(* Logix 5000 project; controller MV vendor 1 type 14 code 217 rev 31.11; software revision 31.00; part 23 of 53 *)
(* tags used below, declared in another part *)
   CheckTimeMask : INT;
   CWD : CHECKWORD_FLAGS;
   Delphi_Does_Eng_Func : BOOL;
   MC_CIP_AV01 : PlantItem;   // CIP_AV01
   MC_CIP_AV02 : PlantItem;   // CIP_AV02
   MC_CIP_AV05 : PlantItem;   // CIP_AV05
   MC_CIP_AV06 : PlantItem;   // CIP_AV06
   MC_CIP_AV07 : PlantItem;   // CIP_AV07
   MC_CIP_AV08 : PlantItem;   // CIP_AV08
   MC_CIP_AV09 : PlantItem;   // CIP_AV09
   MC_CIP_AV10 : PlantItem;   // CIP_AV10
   MC_N255 : INT[255];   // CHECKWORDS Plant item checkword s
   MC_R3R_DR : PlantItem;   // R3R_DR
   MC_R3S_DR : PlantItem;   // R3S_DR
   MC_R3V1 : PlantItem;   // R3V1
   MC_R3V2 : PlantItem;   // R3V2
   MC_SPV5 : PlantItem;   // SPV5
   TempChecktime : DINT;
(* MC_Common, continued *)

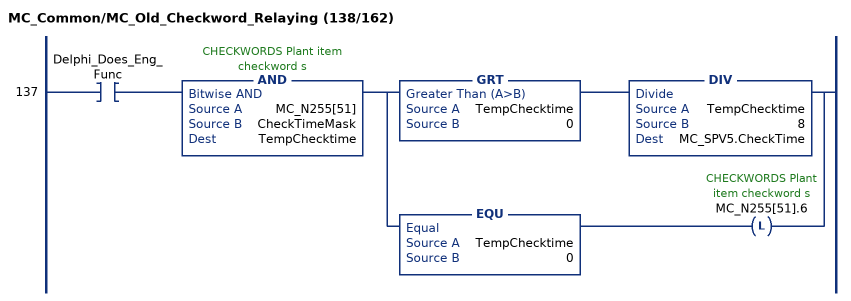
   [picture p410: MC_Common/MC_Old_Checkword_Relaying rungs 137-137]
   137: XIC(Delphi_Does_Eng_Func)AND(MC_N255[51],CheckTimeMask,TempChecktime)[GRT(TempChecktime,0) DIV(TempChecktime,8,MC_SPV5.CheckTime) ,EQU(TempChecktime,0) OTL(MC_N255[51].6) ];
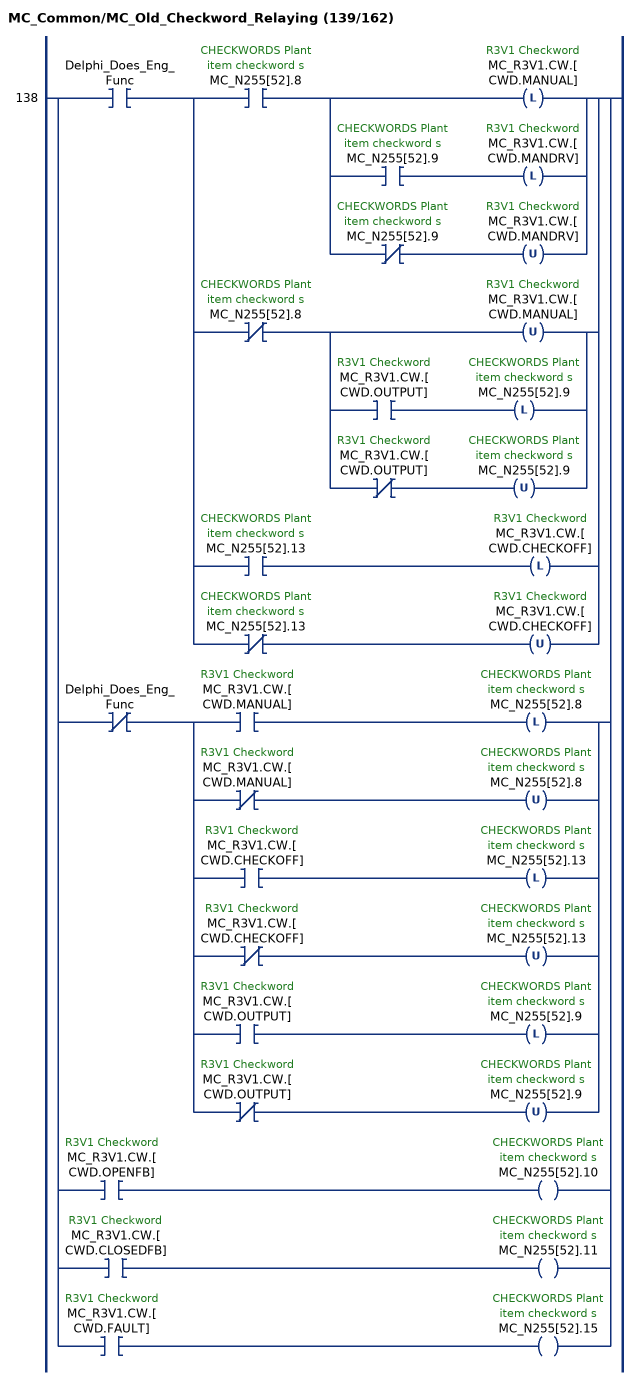
   138: [XIC(Delphi_Does_Eng_Func) [[XIC(MC_N255[52].8) [OTL(MC_R3V1.CW.[CWD.MANUAL]) ,XIC(MC_N255[52].9) OTL(MC_R3V1.CW.[CWD.MANDRV]) ,XIO(MC_N255[52].9) OTU(MC_R3V1.CW.[CWD.MANDRV]) ] ,XIO(MC_N255[52].8) [OTU(MC_R3V1.CW.[CWD.MANUAL]) ,[XIC(MC_R3V1.CW.[CWD.OUTPUT]) OTL(MC_N255[52].9) ,XIO(MC_R3V1.CW.[CWD.OUTPUT]) OTU(MC_N255[52].9) ] ] ] ,[XIC(MC_N255[52].13) OTL(MC_R3V1.CW.[CWD.CHECKOFF]) ,XIO(MC_N255[52].13) OTU(MC_R3V1.CW.[CWD.CHECKOFF]) ] ] ,XIO(Delphi_Does_Eng_Func) [[XIC(MC_R3V1.CW.[CWD.MANUAL]) OTL(MC_N255[52].8) ,XIO(MC_R3V1.CW.[CWD.MANUAL]) OTU(MC_N255[52].8) ] ,[XIC(MC_R3V1.CW.[CWD.CHECKOFF]) OTL(MC_N255[52].13) ,XIO(MC_R3V1.CW.[CWD.CHECKOFF]) OTU(MC_N255[52].13) ] ,[XIC(MC_R3V1.CW.[CWD.OUTPUT]) OTL(MC_N255[52].9) ,XIO(MC_R3V1.CW.[CWD.OUTPUT]) OTU(MC_N255[52].9) ] ] ,XIC(MC_R3V1.CW.[CWD.OPENFB]) OTE(MC_N255[52].10) ,XIC(MC_R3V1.CW.[CWD.CLOSEDFB]) OTE(MC_N255[52].11) ,XIC(MC_R3V1.CW.[CWD.FAULT]) OTE(MC_N255[52].15) ];
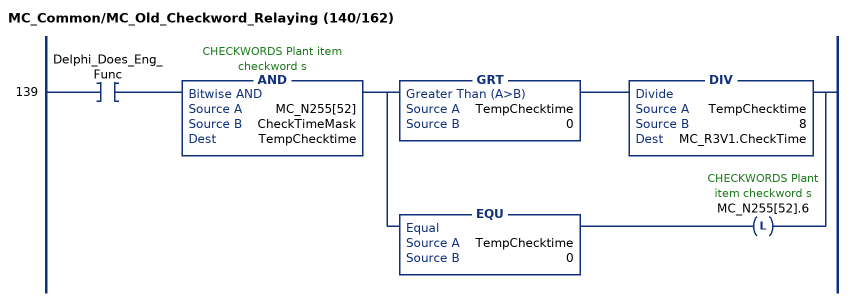
   139: XIC(Delphi_Does_Eng_Func)AND(MC_N255[52],CheckTimeMask,TempChecktime)[GRT(TempChecktime,0) DIV(TempChecktime,8,MC_R3V1.CheckTime) ,EQU(TempChecktime,0) OTL(MC_N255[52].6) ];
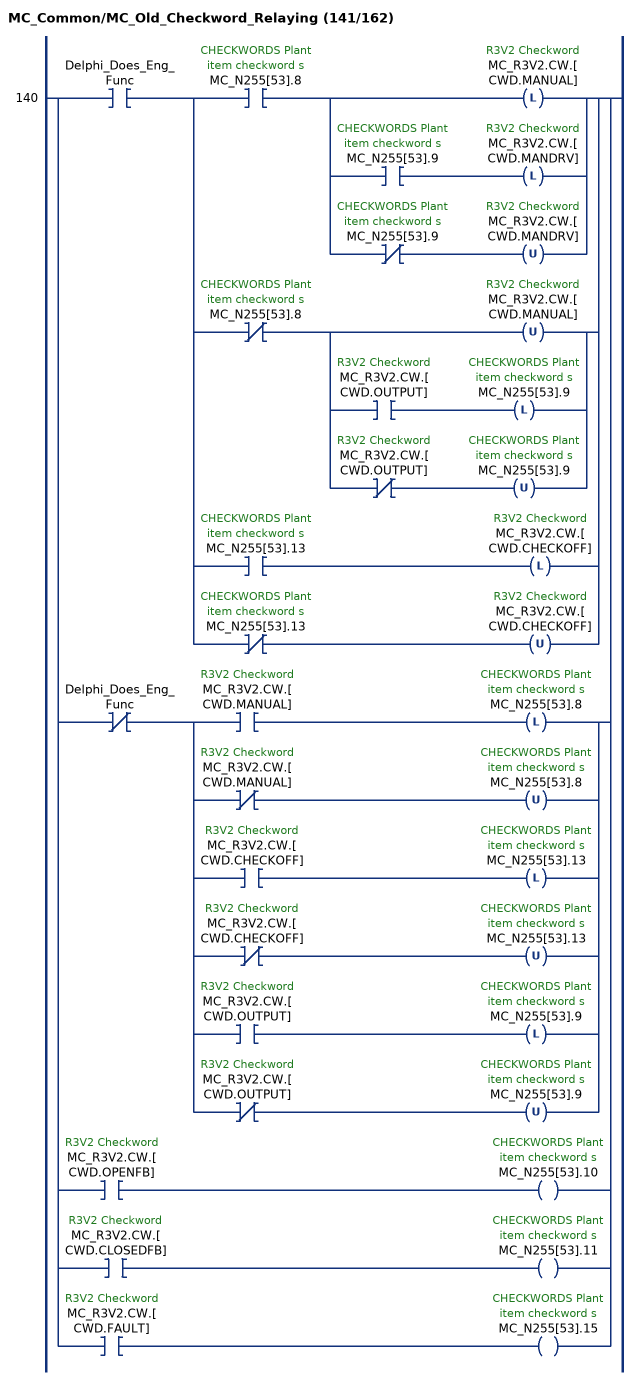
   140: [XIC(Delphi_Does_Eng_Func) [[XIC(MC_N255[53].8) [OTL(MC_R3V2.CW.[CWD.MANUAL]) ,XIC(MC_N255[53].9) OTL(MC_R3V2.CW.[CWD.MANDRV]) ,XIO(MC_N255[53].9) OTU(MC_R3V2.CW.[CWD.MANDRV]) ] ,XIO(MC_N255[53].8) [OTU(MC_R3V2.CW.[CWD.MANUAL]) ,[XIC(MC_R3V2.CW.[CWD.OUTPUT]) OTL(MC_N255[53].9) ,XIO(MC_R3V2.CW.[CWD.OUTPUT]) OTU(MC_N255[53].9) ] ] ] ,[XIC(MC_N255[53].13) OTL(MC_R3V2.CW.[CWD.CHECKOFF]) ,XIO(MC_N255[53].13) OTU(MC_R3V2.CW.[CWD.CHECKOFF]) ] ] ,XIO(Delphi_Does_Eng_Func) [[XIC(MC_R3V2.CW.[CWD.MANUAL]) OTL(MC_N255[53].8) ,XIO(MC_R3V2.CW.[CWD.MANUAL]) OTU(MC_N255[53].8) ] ,[XIC(MC_R3V2.CW.[CWD.CHECKOFF]) OTL(MC_N255[53].13) ,XIO(MC_R3V2.CW.[CWD.CHECKOFF]) OTU(MC_N255[53].13) ] ,[XIC(MC_R3V2.CW.[CWD.OUTPUT]) OTL(MC_N255[53].9) ,XIO(MC_R3V2.CW.[CWD.OUTPUT]) OTU(MC_N255[53].9) ] ] ,XIC(MC_R3V2.CW.[CWD.OPENFB]) OTE(MC_N255[53].10) ,XIC(MC_R3V2.CW.[CWD.CLOSEDFB]) OTE(MC_N255[53].11) ,XIC(MC_R3V2.CW.[CWD.FAULT]) OTE(MC_N255[53].15) ];
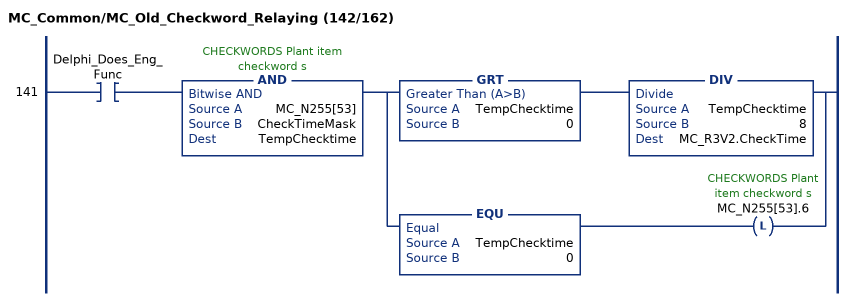
   141: XIC(Delphi_Does_Eng_Func)AND(MC_N255[53],CheckTimeMask,TempChecktime)[GRT(TempChecktime,0) DIV(TempChecktime,8,MC_R3V2.CheckTime) ,EQU(TempChecktime,0) OTL(MC_N255[53].6) ];
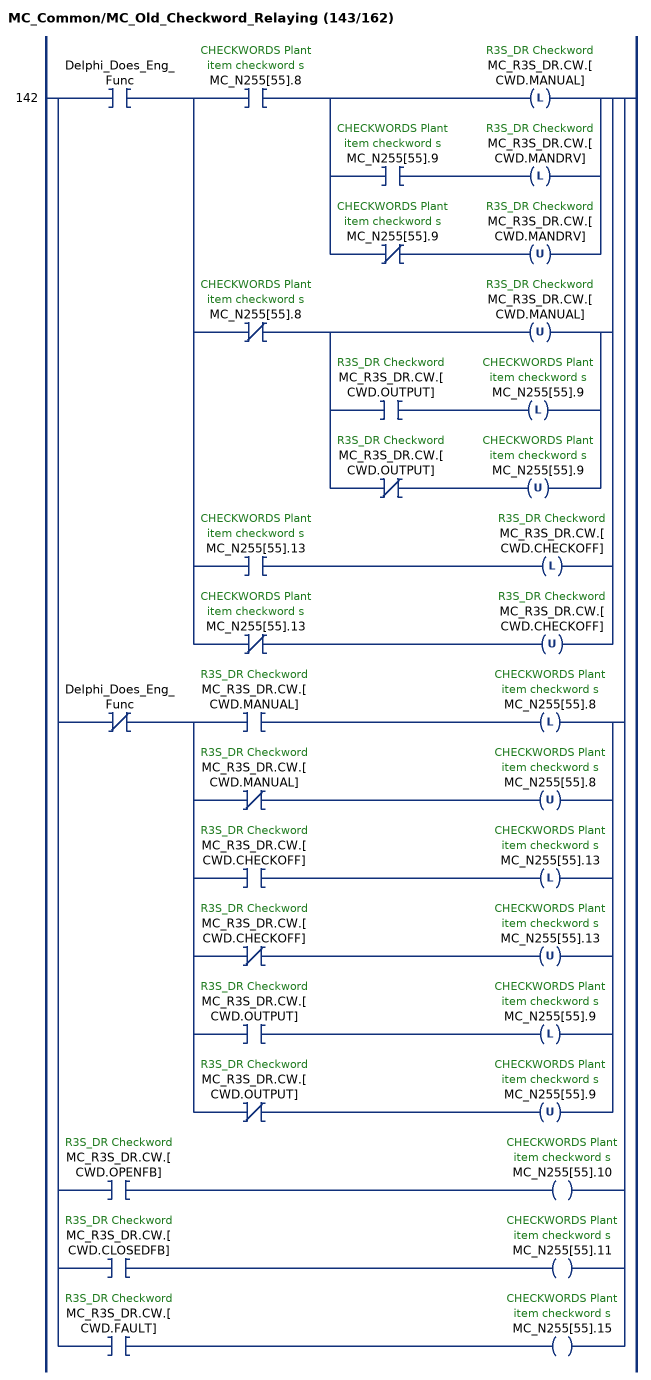
   142: [XIC(Delphi_Does_Eng_Func) [[XIC(MC_N255[55].8) [OTL(MC_R3S_DR.CW.[CWD.MANUAL]) ,XIC(MC_N255[55].9) OTL(MC_R3S_DR.CW.[CWD.MANDRV]) ,XIO(MC_N255[55].9) OTU(MC_R3S_DR.CW.[CWD.MANDRV]) ] ,XIO(MC_N255[55].8) [OTU(MC_R3S_DR.CW.[CWD.MANUAL]) ,[XIC(MC_R3S_DR.CW.[CWD.OUTPUT]) OTL(MC_N255[55].9) ,XIO(MC_R3S_DR.CW.[CWD.OUTPUT]) OTU(MC_N255[55].9) ] ] ] ,[XIC(MC_N255[55].13) OTL(MC_R3S_DR.CW.[CWD.CHECKOFF]) ,XIO(MC_N255[55].13) OTU(MC_R3S_DR.CW.[CWD.CHECKOFF]) ] ] ,XIO(Delphi_Does_Eng_Func) [[XIC(MC_R3S_DR.CW.[CWD.MANUAL]) OTL(MC_N255[55].8) ,XIO(MC_R3S_DR.CW.[CWD.MANUAL]) OTU(MC_N255[55].8) ] ,[XIC(MC_R3S_DR.CW.[CWD.CHECKOFF]) OTL(MC_N255[55].13) ,XIO(MC_R3S_DR.CW.[CWD.CHECKOFF]) OTU(MC_N255[55].13) ] ,[XIC(MC_R3S_DR.CW.[CWD.OUTPUT]) OTL(MC_N255[55].9) ,XIO(MC_R3S_DR.CW.[CWD.OUTPUT]) OTU(MC_N255[55].9) ] ] ,XIC(MC_R3S_DR.CW.[CWD.OPENFB]) OTE(MC_N255[55].10) ,XIC(MC_R3S_DR.CW.[CWD.CLOSEDFB]) OTE(MC_N255[55].11) ,XIC(MC_R3S_DR.CW.[CWD.FAULT]) OTE(MC_N255[55].15) ];
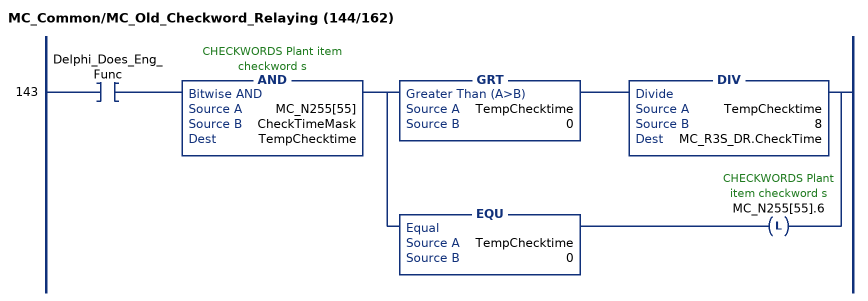
   143: XIC(Delphi_Does_Eng_Func)AND(MC_N255[55],CheckTimeMask,TempChecktime)[GRT(TempChecktime,0) DIV(TempChecktime,8,MC_R3S_DR.CheckTime) ,EQU(TempChecktime,0) OTL(MC_N255[55].6) ];
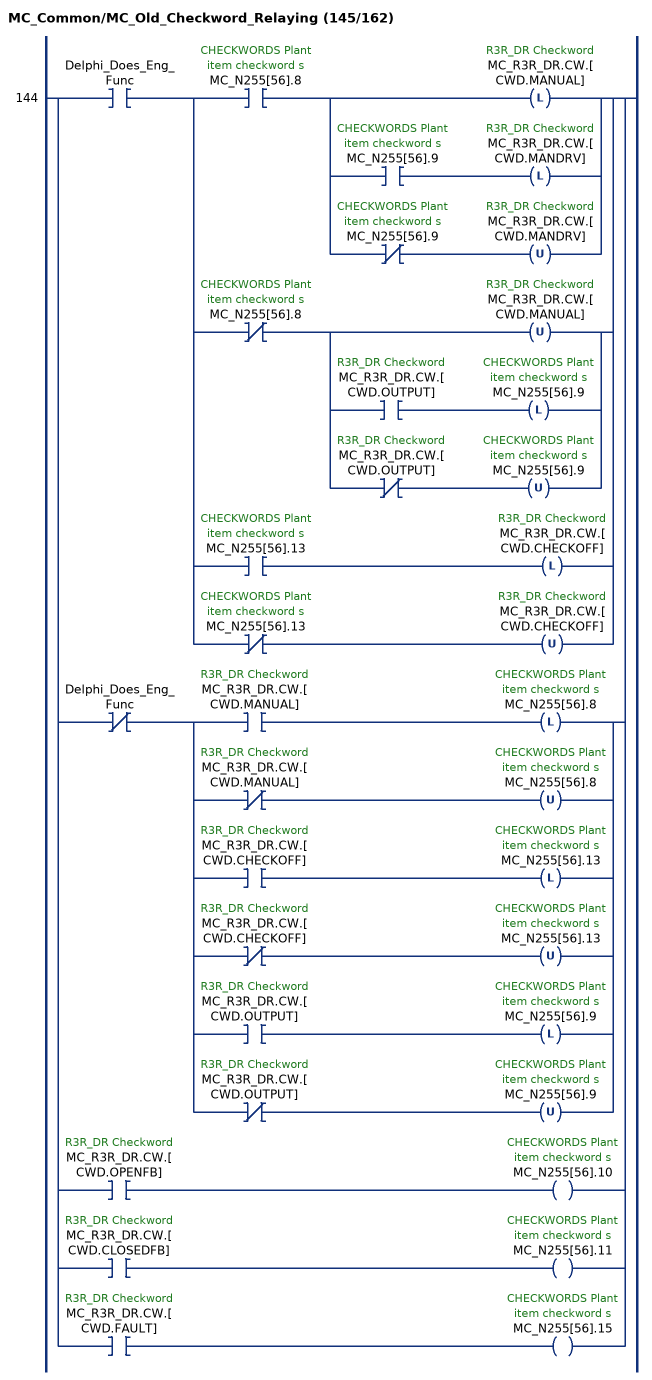
   144: [XIC(Delphi_Does_Eng_Func) [[XIC(MC_N255[56].8) [OTL(MC_R3R_DR.CW.[CWD.MANUAL]) ,XIC(MC_N255[56].9) OTL(MC_R3R_DR.CW.[CWD.MANDRV]) ,XIO(MC_N255[56].9) OTU(MC_R3R_DR.CW.[CWD.MANDRV]) ] ,XIO(MC_N255[56].8) [OTU(MC_R3R_DR.CW.[CWD.MANUAL]) ,[XIC(MC_R3R_DR.CW.[CWD.OUTPUT]) OTL(MC_N255[56].9) ,XIO(MC_R3R_DR.CW.[CWD.OUTPUT]) OTU(MC_N255[56].9) ] ] ] ,[XIC(MC_N255[56].13) OTL(MC_R3R_DR.CW.[CWD.CHECKOFF]) ,XIO(MC_N255[56].13) OTU(MC_R3R_DR.CW.[CWD.CHECKOFF]) ] ] ,XIO(Delphi_Does_Eng_Func) [[XIC(MC_R3R_DR.CW.[CWD.MANUAL]) OTL(MC_N255[56].8) ,XIO(MC_R3R_DR.CW.[CWD.MANUAL]) OTU(MC_N255[56].8) ] ,[XIC(MC_R3R_DR.CW.[CWD.CHECKOFF]) OTL(MC_N255[56].13) ,XIO(MC_R3R_DR.CW.[CWD.CHECKOFF]) OTU(MC_N255[56].13) ] ,[XIC(MC_R3R_DR.CW.[CWD.OUTPUT]) OTL(MC_N255[56].9) ,XIO(MC_R3R_DR.CW.[CWD.OUTPUT]) OTU(MC_N255[56].9) ] ] ,XIC(MC_R3R_DR.CW.[CWD.OPENFB]) OTE(MC_N255[56].10) ,XIC(MC_R3R_DR.CW.[CWD.CLOSEDFB]) OTE(MC_N255[56].11) ,XIC(MC_R3R_DR.CW.[CWD.FAULT]) OTE(MC_N255[56].15) ];
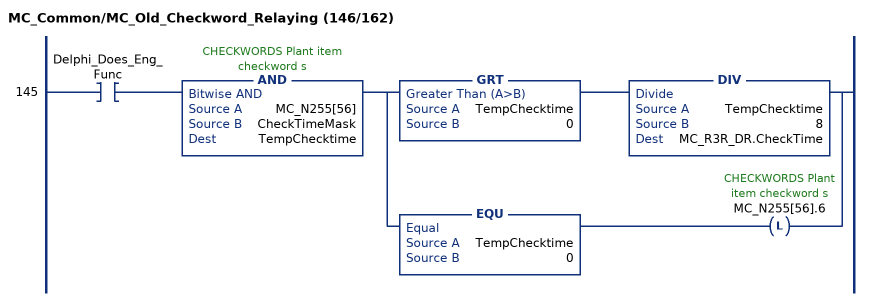
   145: XIC(Delphi_Does_Eng_Func)AND(MC_N255[56],CheckTimeMask,TempChecktime)[GRT(TempChecktime,0) DIV(TempChecktime,8,MC_R3R_DR.CheckTime) ,EQU(TempChecktime,0) OTL(MC_N255[56].6) ];
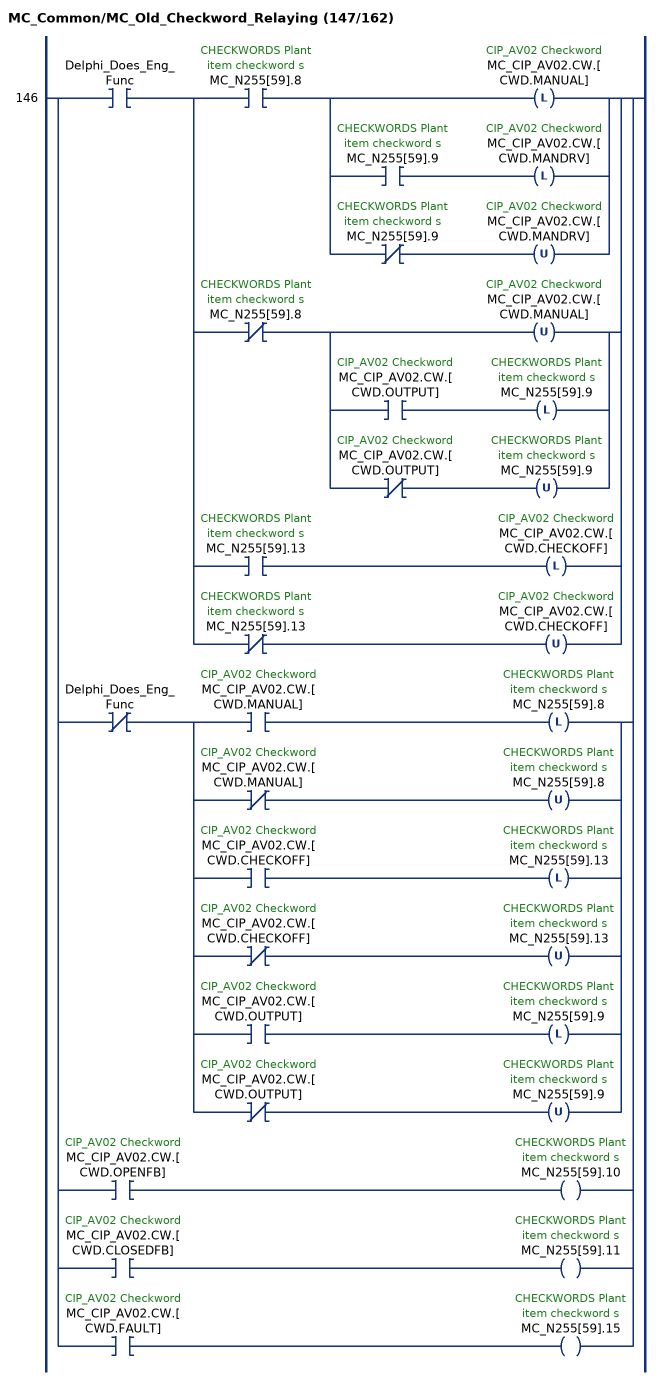
   146: [XIC(Delphi_Does_Eng_Func) [[XIC(MC_N255[59].8) [OTL(MC_CIP_AV02.CW.[CWD.MANUAL]) ,XIC(MC_N255[59].9) OTL(MC_CIP_AV02.CW.[CWD.MANDRV]) ,XIO(MC_N255[59].9) OTU(MC_CIP_AV02.CW.[CWD.MANDRV]) ] ,XIO(MC_N255[59].8) [OTU(MC_CIP_AV02.CW.[CWD.MANUAL]) ,[XIC(MC_CIP_AV02.CW.[CWD.OUTPUT]) OTL(MC_N255[59].9) ,XIO(MC_CIP_AV02.CW.[CWD.OUTPUT]) OTU(MC_N255[59].9) ] ] ] ,[XIC(MC_N255[59].13) OTL(MC_CIP_AV02.CW.[CWD.CHECKOFF]) ,XIO(MC_N255[59].13) OTU(MC_CIP_AV02.CW.[CWD.CHECKOFF]) ] ] ,XIO(Delphi_Does_Eng_Func) [[XIC(MC_CIP_AV02.CW.[CWD.MANUAL]) OTL(MC_N255[59].8) ,XIO(MC_CIP_AV02.CW.[CWD.MANUAL]) OTU(MC_N255[59].8) ] ,[XIC(MC_CIP_AV02.CW.[CWD.CHECKOFF]) OTL(MC_N255[59].13) ,XIO(MC_CIP_AV02.CW.[CWD.CHECKOFF]) OTU(MC_N255[59].13) ] ,[XIC(MC_CIP_AV02.CW.[CWD.OUTPUT]) OTL(MC_N255[59].9) ,XIO(MC_CIP_AV02.CW.[CWD.OUTPUT]) OTU(MC_N255[59].9) ] ] ,XIC(MC_CIP_AV02.CW.[CWD.OPENFB]) OTE(MC_N255[59].10) ,XIC(MC_CIP_AV02.CW.[CWD.CLOSEDFB]) OTE(MC_N255[59].11) ,XIC(MC_CIP_AV02.CW.[CWD.FAULT]) OTE(MC_N255[59].15) ];
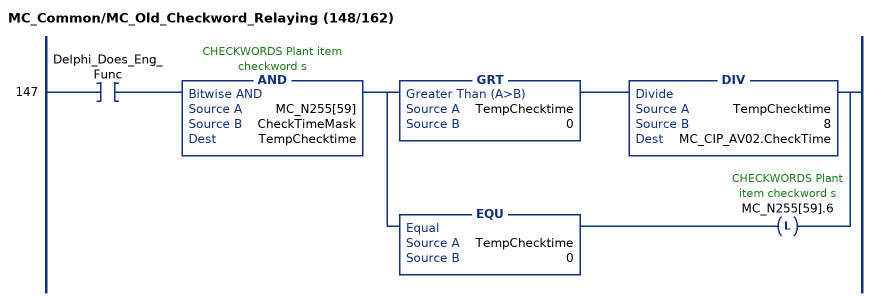
   147: XIC(Delphi_Does_Eng_Func)AND(MC_N255[59],CheckTimeMask,TempChecktime)[GRT(TempChecktime,0) DIV(TempChecktime,8,MC_CIP_AV02.CheckTime) ,EQU(TempChecktime,0) OTL(MC_N255[59].6) ];
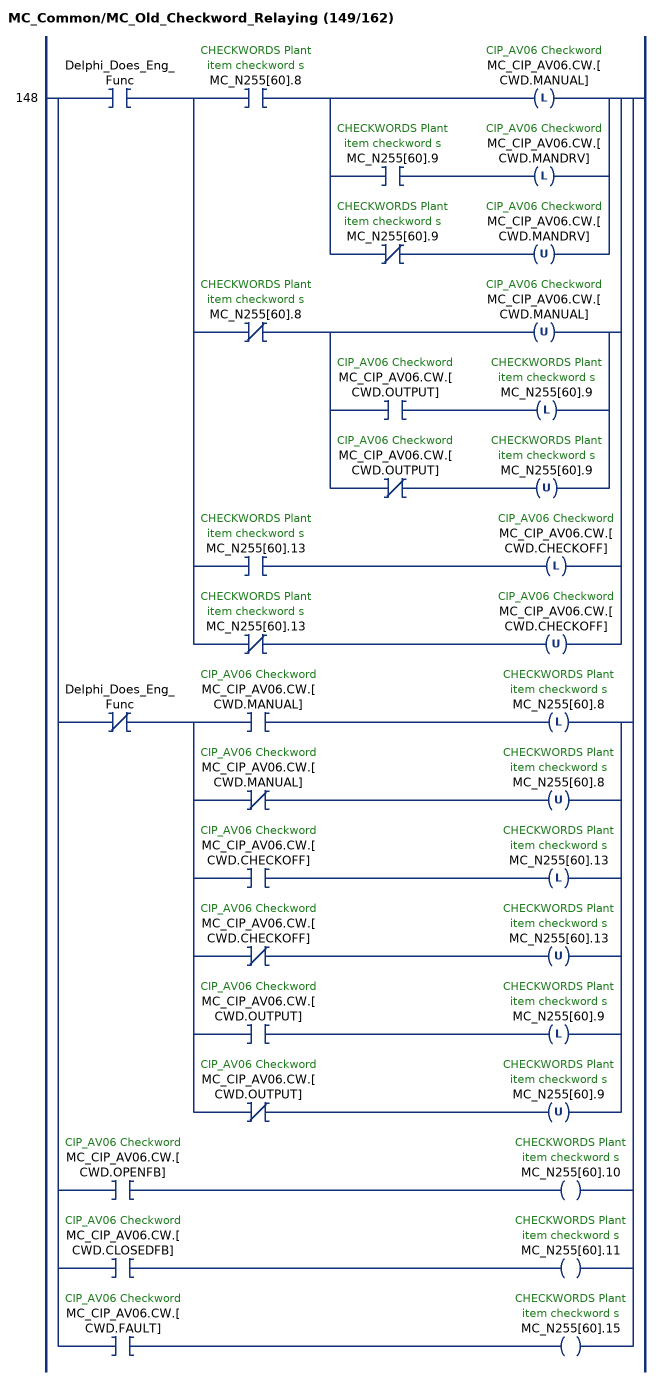
   148: [XIC(Delphi_Does_Eng_Func) [[XIC(MC_N255[60].8) [OTL(MC_CIP_AV06.CW.[CWD.MANUAL]) ,XIC(MC_N255[60].9) OTL(MC_CIP_AV06.CW.[CWD.MANDRV]) ,XIO(MC_N255[60].9) OTU(MC_CIP_AV06.CW.[CWD.MANDRV]) ] ,XIO(MC_N255[60].8) [OTU(MC_CIP_AV06.CW.[CWD.MANUAL]) ,[XIC(MC_CIP_AV06.CW.[CWD.OUTPUT]) OTL(MC_N255[60].9) ,XIO(MC_CIP_AV06.CW.[CWD.OUTPUT]) OTU(MC_N255[60].9) ] ] ] ,[XIC(MC_N255[60].13) OTL(MC_CIP_AV06.CW.[CWD.CHECKOFF]) ,XIO(MC_N255[60].13) OTU(MC_CIP_AV06.CW.[CWD.CHECKOFF]) ] ] ,XIO(Delphi_Does_Eng_Func) [[XIC(MC_CIP_AV06.CW.[CWD.MANUAL]) OTL(MC_N255[60].8) ,XIO(MC_CIP_AV06.CW.[CWD.MANUAL]) OTU(MC_N255[60].8) ] ,[XIC(MC_CIP_AV06.CW.[CWD.CHECKOFF]) OTL(MC_N255[60].13) ,XIO(MC_CIP_AV06.CW.[CWD.CHECKOFF]) OTU(MC_N255[60].13) ] ,[XIC(MC_CIP_AV06.CW.[CWD.OUTPUT]) OTL(MC_N255[60].9) ,XIO(MC_CIP_AV06.CW.[CWD.OUTPUT]) OTU(MC_N255[60].9) ] ] ,XIC(MC_CIP_AV06.CW.[CWD.OPENFB]) OTE(MC_N255[60].10) ,XIC(MC_CIP_AV06.CW.[CWD.CLOSEDFB]) OTE(MC_N255[60].11) ,XIC(MC_CIP_AV06.CW.[CWD.FAULT]) OTE(MC_N255[60].15) ];
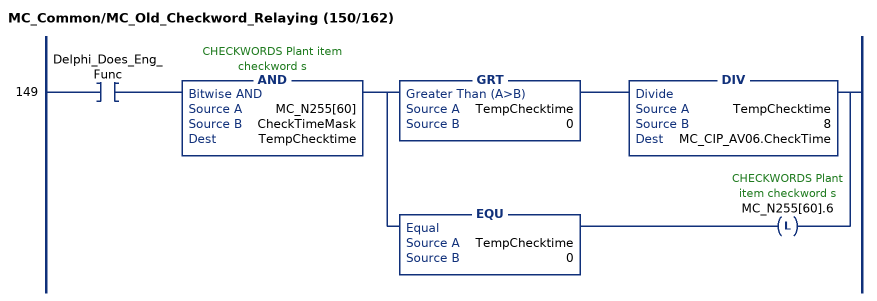
   149: XIC(Delphi_Does_Eng_Func)AND(MC_N255[60],CheckTimeMask,TempChecktime)[GRT(TempChecktime,0) DIV(TempChecktime,8,MC_CIP_AV06.CheckTime) ,EQU(TempChecktime,0) OTL(MC_N255[60].6) ];
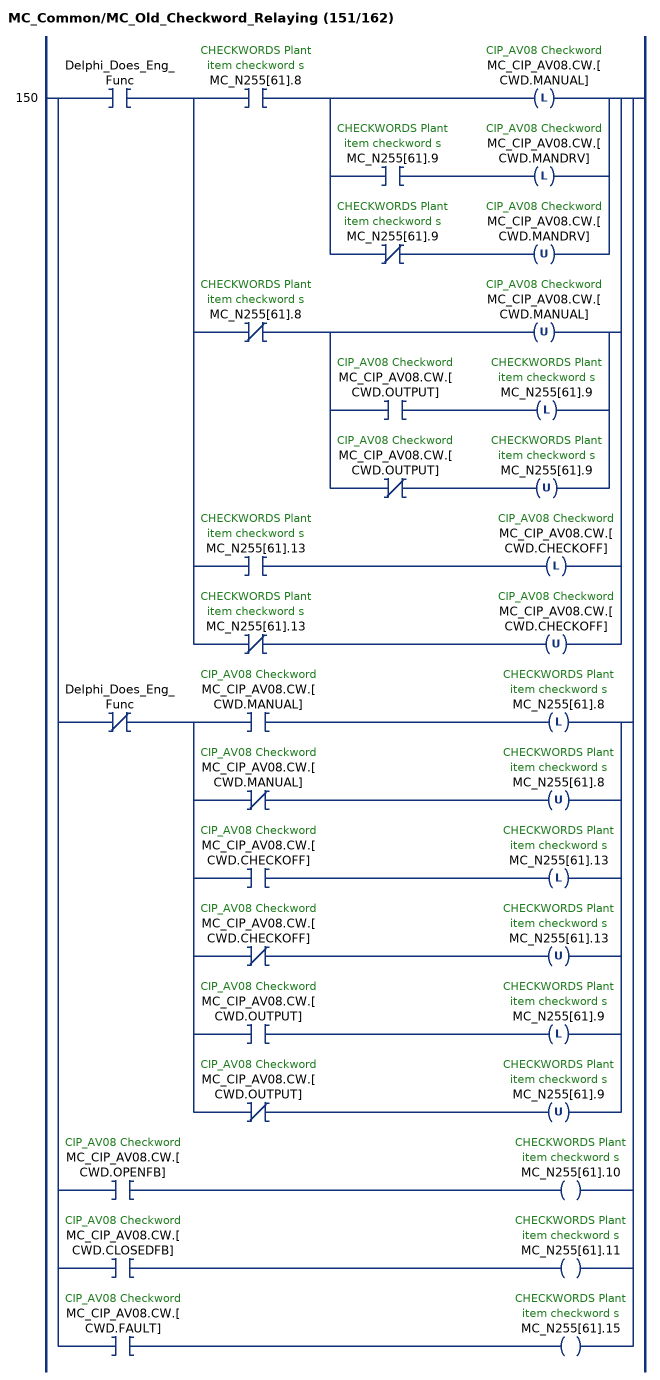
   150: [XIC(Delphi_Does_Eng_Func) [[XIC(MC_N255[61].8) [OTL(MC_CIP_AV08.CW.[CWD.MANUAL]) ,XIC(MC_N255[61].9) OTL(MC_CIP_AV08.CW.[CWD.MANDRV]) ,XIO(MC_N255[61].9) OTU(MC_CIP_AV08.CW.[CWD.MANDRV]) ] ,XIO(MC_N255[61].8) [OTU(MC_CIP_AV08.CW.[CWD.MANUAL]) ,[XIC(MC_CIP_AV08.CW.[CWD.OUTPUT]) OTL(MC_N255[61].9) ,XIO(MC_CIP_AV08.CW.[CWD.OUTPUT]) OTU(MC_N255[61].9) ] ] ] ,[XIC(MC_N255[61].13) OTL(MC_CIP_AV08.CW.[CWD.CHECKOFF]) ,XIO(MC_N255[61].13) OTU(MC_CIP_AV08.CW.[CWD.CHECKOFF]) ] ] ,XIO(Delphi_Does_Eng_Func) [[XIC(MC_CIP_AV08.CW.[CWD.MANUAL]) OTL(MC_N255[61].8) ,XIO(MC_CIP_AV08.CW.[CWD.MANUAL]) OTU(MC_N255[61].8) ] ,[XIC(MC_CIP_AV08.CW.[CWD.CHECKOFF]) OTL(MC_N255[61].13) ,XIO(MC_CIP_AV08.CW.[CWD.CHECKOFF]) OTU(MC_N255[61].13) ] ,[XIC(MC_CIP_AV08.CW.[CWD.OUTPUT]) OTL(MC_N255[61].9) ,XIO(MC_CIP_AV08.CW.[CWD.OUTPUT]) OTU(MC_N255[61].9) ] ] ,XIC(MC_CIP_AV08.CW.[CWD.OPENFB]) OTE(MC_N255[61].10) ,XIC(MC_CIP_AV08.CW.[CWD.CLOSEDFB]) OTE(MC_N255[61].11) ,XIC(MC_CIP_AV08.CW.[CWD.FAULT]) OTE(MC_N255[61].15) ];
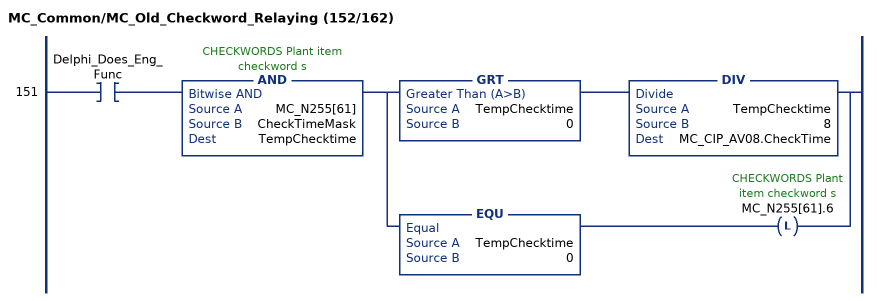
   151: XIC(Delphi_Does_Eng_Func)AND(MC_N255[61],CheckTimeMask,TempChecktime)[GRT(TempChecktime,0) DIV(TempChecktime,8,MC_CIP_AV08.CheckTime) ,EQU(TempChecktime,0) OTL(MC_N255[61].6) ];
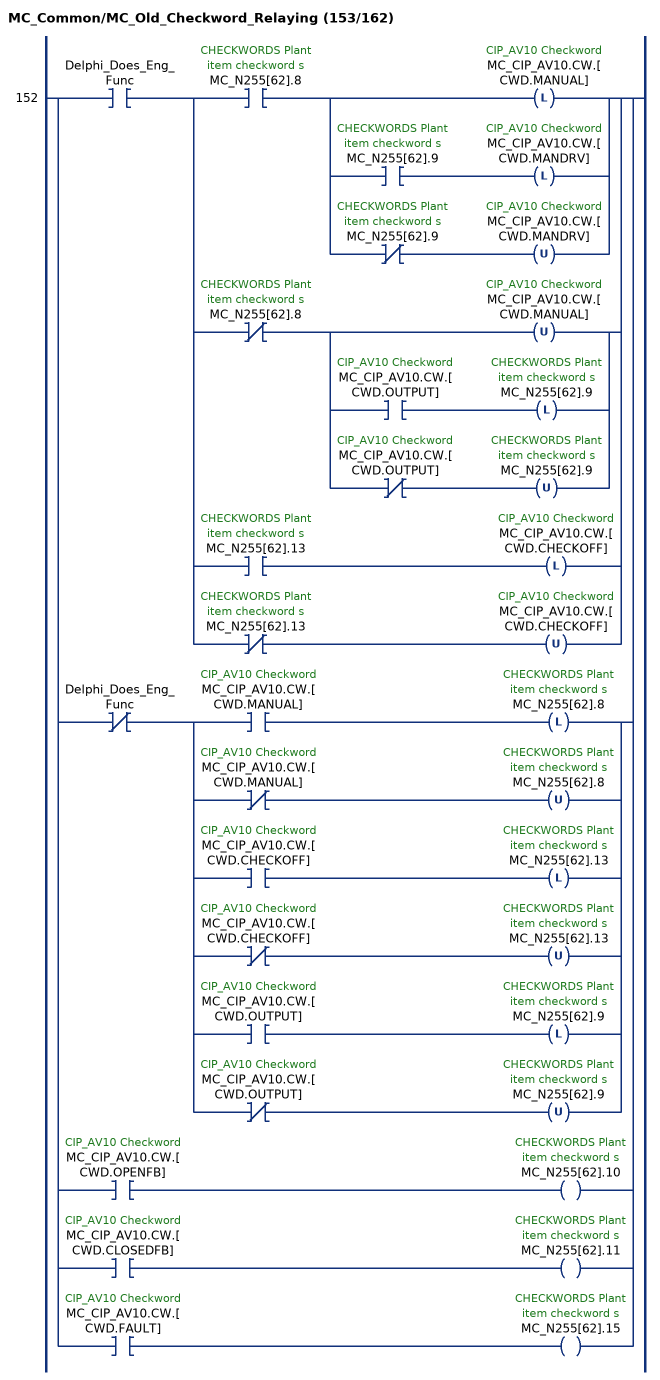
   152: [XIC(Delphi_Does_Eng_Func) [[XIC(MC_N255[62].8) [OTL(MC_CIP_AV10.CW.[CWD.MANUAL]) ,XIC(MC_N255[62].9) OTL(MC_CIP_AV10.CW.[CWD.MANDRV]) ,XIO(MC_N255[62].9) OTU(MC_CIP_AV10.CW.[CWD.MANDRV]) ] ,XIO(MC_N255[62].8) [OTU(MC_CIP_AV10.CW.[CWD.MANUAL]) ,[XIC(MC_CIP_AV10.CW.[CWD.OUTPUT]) OTL(MC_N255[62].9) ,XIO(MC_CIP_AV10.CW.[CWD.OUTPUT]) OTU(MC_N255[62].9) ] ] ] ,[XIC(MC_N255[62].13) OTL(MC_CIP_AV10.CW.[CWD.CHECKOFF]) ,XIO(MC_N255[62].13) OTU(MC_CIP_AV10.CW.[CWD.CHECKOFF]) ] ] ,XIO(Delphi_Does_Eng_Func) [[XIC(MC_CIP_AV10.CW.[CWD.MANUAL]) OTL(MC_N255[62].8) ,XIO(MC_CIP_AV10.CW.[CWD.MANUAL]) OTU(MC_N255[62].8) ] ,[XIC(MC_CIP_AV10.CW.[CWD.CHECKOFF]) OTL(MC_N255[62].13) ,XIO(MC_CIP_AV10.CW.[CWD.CHECKOFF]) OTU(MC_N255[62].13) ] ,[XIC(MC_CIP_AV10.CW.[CWD.OUTPUT]) OTL(MC_N255[62].9) ,XIO(MC_CIP_AV10.CW.[CWD.OUTPUT]) OTU(MC_N255[62].9) ] ] ,XIC(MC_CIP_AV10.CW.[CWD.OPENFB]) OTE(MC_N255[62].10) ,XIC(MC_CIP_AV10.CW.[CWD.CLOSEDFB]) OTE(MC_N255[62].11) ,XIC(MC_CIP_AV10.CW.[CWD.FAULT]) OTE(MC_N255[62].15) ];
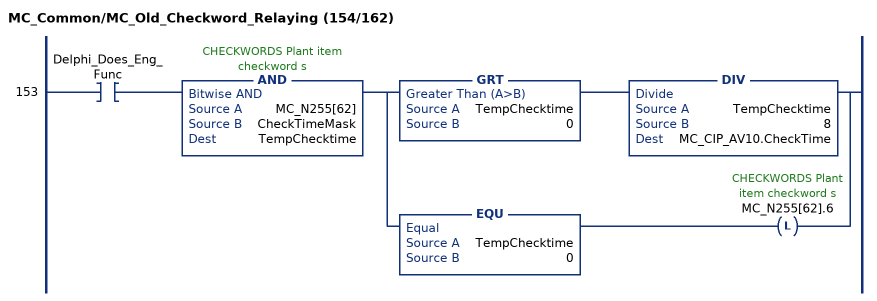
   153: XIC(Delphi_Does_Eng_Func)AND(MC_N255[62],CheckTimeMask,TempChecktime)[GRT(TempChecktime,0) DIV(TempChecktime,8,MC_CIP_AV10.CheckTime) ,EQU(TempChecktime,0) OTL(MC_N255[62].6) ];
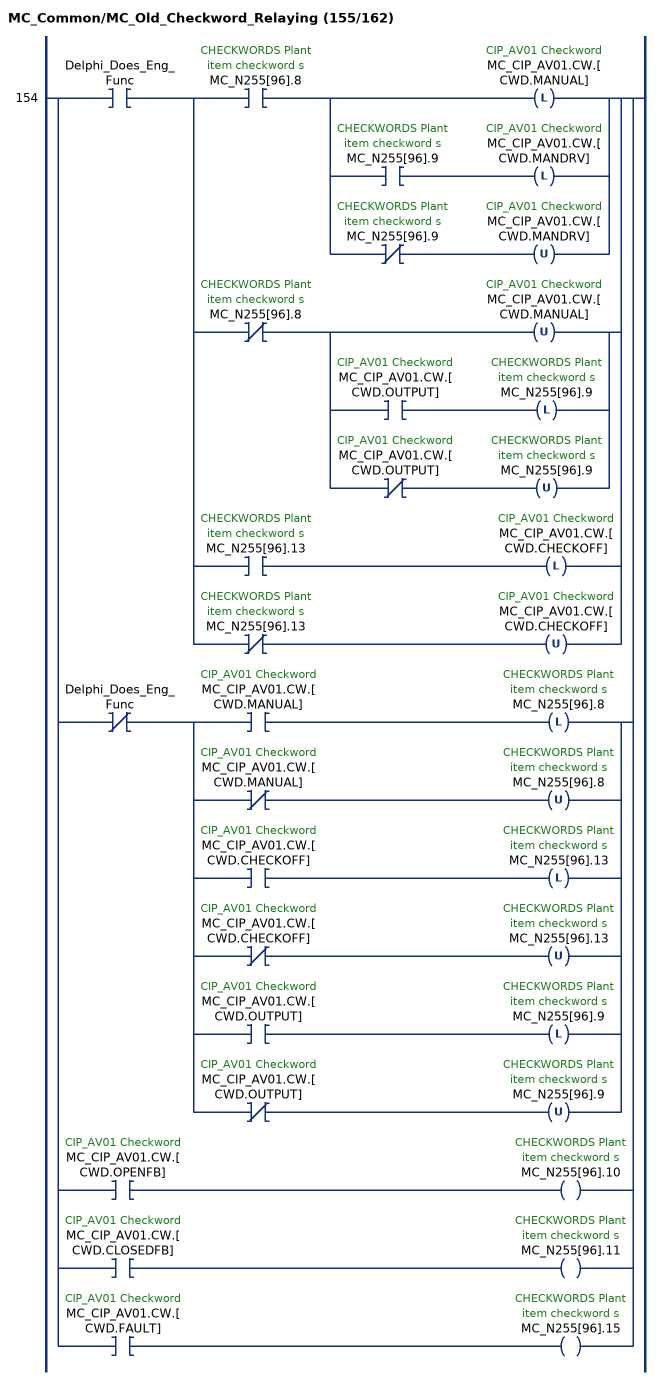
   154: [XIC(Delphi_Does_Eng_Func) [[XIC(MC_N255[96].8) [OTL(MC_CIP_AV01.CW.[CWD.MANUAL]) ,XIC(MC_N255[96].9) OTL(MC_CIP_AV01.CW.[CWD.MANDRV]) ,XIO(MC_N255[96].9) OTU(MC_CIP_AV01.CW.[CWD.MANDRV]) ] ,XIO(MC_N255[96].8) [OTU(MC_CIP_AV01.CW.[CWD.MANUAL]) ,[XIC(MC_CIP_AV01.CW.[CWD.OUTPUT]) OTL(MC_N255[96].9) ,XIO(MC_CIP_AV01.CW.[CWD.OUTPUT]) OTU(MC_N255[96].9) ] ] ] ,[XIC(MC_N255[96].13) OTL(MC_CIP_AV01.CW.[CWD.CHECKOFF]) ,XIO(MC_N255[96].13) OTU(MC_CIP_AV01.CW.[CWD.CHECKOFF]) ] ] ,XIO(Delphi_Does_Eng_Func) [[XIC(MC_CIP_AV01.CW.[CWD.MANUAL]) OTL(MC_N255[96].8) ,XIO(MC_CIP_AV01.CW.[CWD.MANUAL]) OTU(MC_N255[96].8) ] ,[XIC(MC_CIP_AV01.CW.[CWD.CHECKOFF]) OTL(MC_N255[96].13) ,XIO(MC_CIP_AV01.CW.[CWD.CHECKOFF]) OTU(MC_N255[96].13) ] ,[XIC(MC_CIP_AV01.CW.[CWD.OUTPUT]) OTL(MC_N255[96].9) ,XIO(MC_CIP_AV01.CW.[CWD.OUTPUT]) OTU(MC_N255[96].9) ] ] ,XIC(MC_CIP_AV01.CW.[CWD.OPENFB]) OTE(MC_N255[96].10) ,XIC(MC_CIP_AV01.CW.[CWD.CLOSEDFB]) OTE(MC_N255[96].11) ,XIC(MC_CIP_AV01.CW.[CWD.FAULT]) OTE(MC_N255[96].15) ];
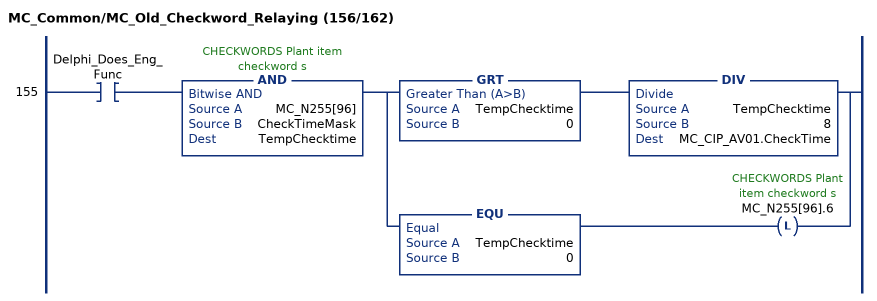
   155: XIC(Delphi_Does_Eng_Func)AND(MC_N255[96],CheckTimeMask,TempChecktime)[GRT(TempChecktime,0) DIV(TempChecktime,8,MC_CIP_AV01.CheckTime) ,EQU(TempChecktime,0) OTL(MC_N255[96].6) ];
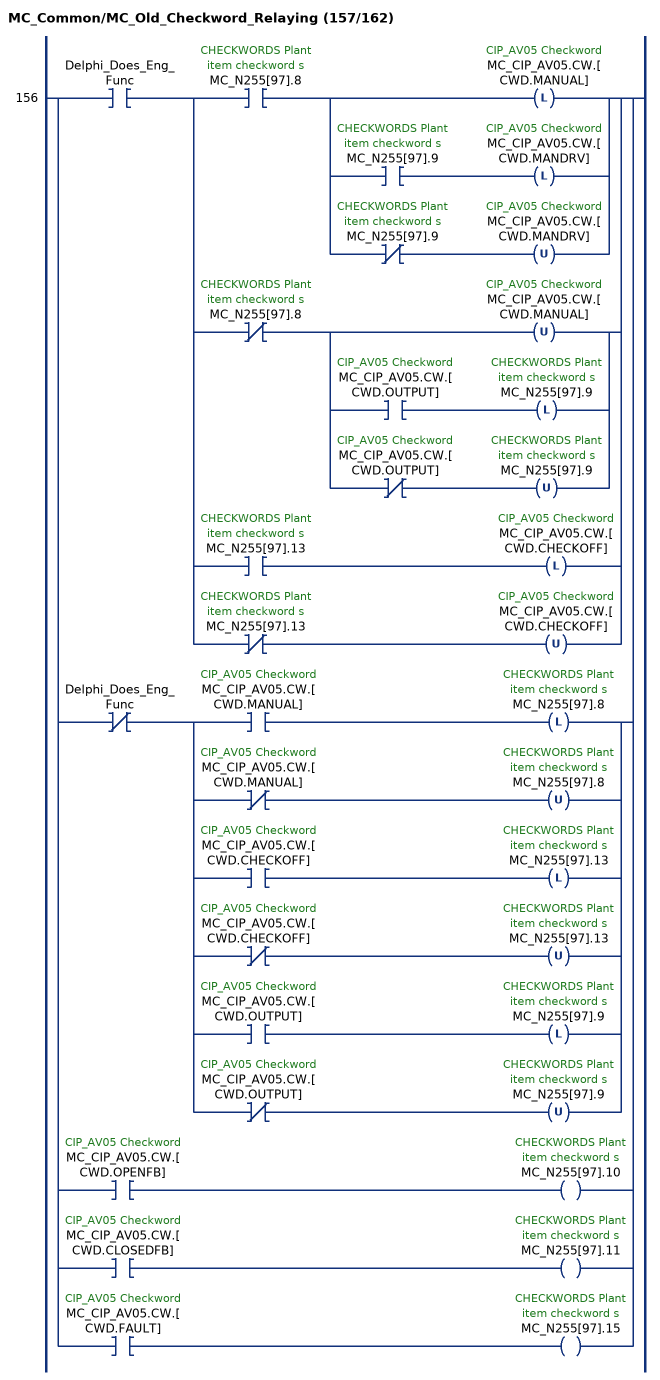
   156: [XIC(Delphi_Does_Eng_Func) [[XIC(MC_N255[97].8) [OTL(MC_CIP_AV05.CW.[CWD.MANUAL]) ,XIC(MC_N255[97].9) OTL(MC_CIP_AV05.CW.[CWD.MANDRV]) ,XIO(MC_N255[97].9) OTU(MC_CIP_AV05.CW.[CWD.MANDRV]) ] ,XIO(MC_N255[97].8) [OTU(MC_CIP_AV05.CW.[CWD.MANUAL]) ,[XIC(MC_CIP_AV05.CW.[CWD.OUTPUT]) OTL(MC_N255[97].9) ,XIO(MC_CIP_AV05.CW.[CWD.OUTPUT]) OTU(MC_N255[97].9) ] ] ] ,[XIC(MC_N255[97].13) OTL(MC_CIP_AV05.CW.[CWD.CHECKOFF]) ,XIO(MC_N255[97].13) OTU(MC_CIP_AV05.CW.[CWD.CHECKOFF]) ] ] ,XIO(Delphi_Does_Eng_Func) [[XIC(MC_CIP_AV05.CW.[CWD.MANUAL]) OTL(MC_N255[97].8) ,XIO(MC_CIP_AV05.CW.[CWD.MANUAL]) OTU(MC_N255[97].8) ] ,[XIC(MC_CIP_AV05.CW.[CWD.CHECKOFF]) OTL(MC_N255[97].13) ,XIO(MC_CIP_AV05.CW.[CWD.CHECKOFF]) OTU(MC_N255[97].13) ] ,[XIC(MC_CIP_AV05.CW.[CWD.OUTPUT]) OTL(MC_N255[97].9) ,XIO(MC_CIP_AV05.CW.[CWD.OUTPUT]) OTU(MC_N255[97].9) ] ] ,XIC(MC_CIP_AV05.CW.[CWD.OPENFB]) OTE(MC_N255[97].10) ,XIC(MC_CIP_AV05.CW.[CWD.CLOSEDFB]) OTE(MC_N255[97].11) ,XIC(MC_CIP_AV05.CW.[CWD.FAULT]) OTE(MC_N255[97].15) ];
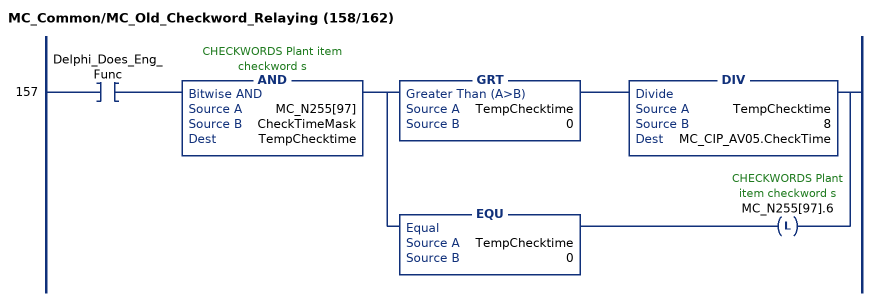
   157: XIC(Delphi_Does_Eng_Func)AND(MC_N255[97],CheckTimeMask,TempChecktime)[GRT(TempChecktime,0) DIV(TempChecktime,8,MC_CIP_AV05.CheckTime) ,EQU(TempChecktime,0) OTL(MC_N255[97].6) ];
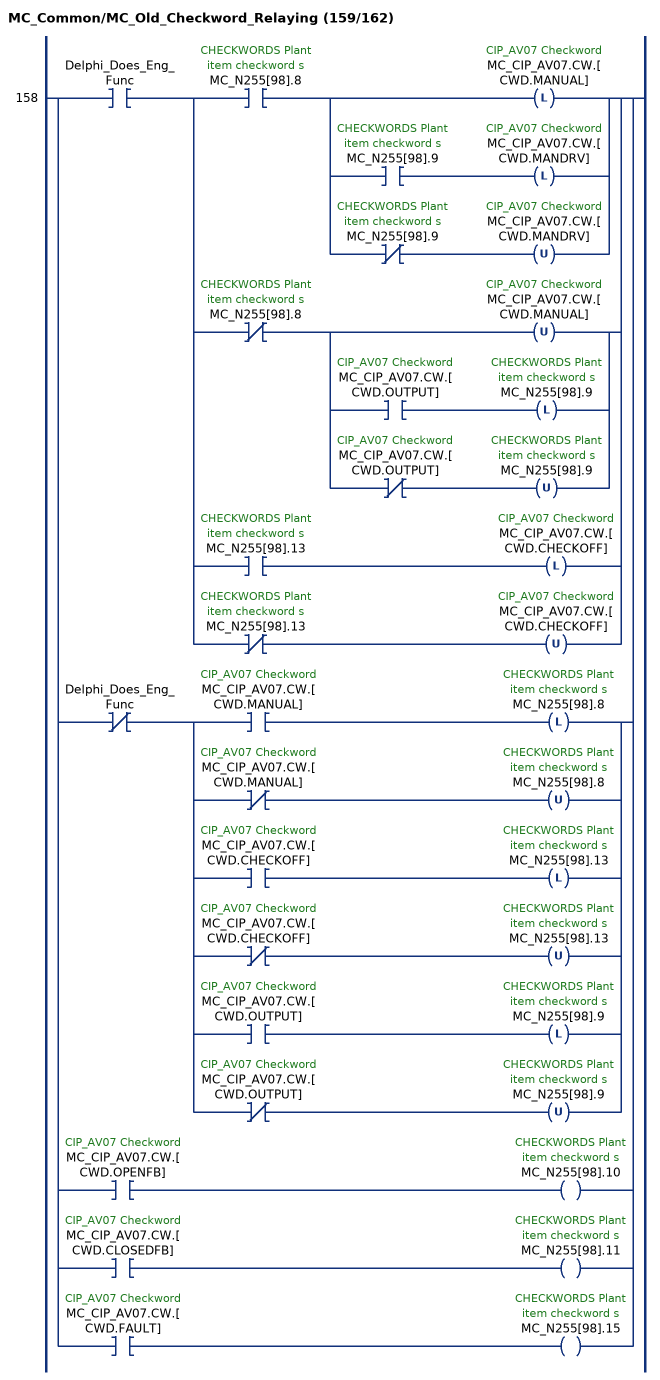
   158: [XIC(Delphi_Does_Eng_Func) [[XIC(MC_N255[98].8) [OTL(MC_CIP_AV07.CW.[CWD.MANUAL]) ,XIC(MC_N255[98].9) OTL(MC_CIP_AV07.CW.[CWD.MANDRV]) ,XIO(MC_N255[98].9) OTU(MC_CIP_AV07.CW.[CWD.MANDRV]) ] ,XIO(MC_N255[98].8) [OTU(MC_CIP_AV07.CW.[CWD.MANUAL]) ,[XIC(MC_CIP_AV07.CW.[CWD.OUTPUT]) OTL(MC_N255[98].9) ,XIO(MC_CIP_AV07.CW.[CWD.OUTPUT]) OTU(MC_N255[98].9) ] ] ] ,[XIC(MC_N255[98].13) OTL(MC_CIP_AV07.CW.[CWD.CHECKOFF]) ,XIO(MC_N255[98].13) OTU(MC_CIP_AV07.CW.[CWD.CHECKOFF]) ] ] ,XIO(Delphi_Does_Eng_Func) [[XIC(MC_CIP_AV07.CW.[CWD.MANUAL]) OTL(MC_N255[98].8) ,XIO(MC_CIP_AV07.CW.[CWD.MANUAL]) OTU(MC_N255[98].8) ] ,[XIC(MC_CIP_AV07.CW.[CWD.CHECKOFF]) OTL(MC_N255[98].13) ,XIO(MC_CIP_AV07.CW.[CWD.CHECKOFF]) OTU(MC_N255[98].13) ] ,[XIC(MC_CIP_AV07.CW.[CWD.OUTPUT]) OTL(MC_N255[98].9) ,XIO(MC_CIP_AV07.CW.[CWD.OUTPUT]) OTU(MC_N255[98].9) ] ] ,XIC(MC_CIP_AV07.CW.[CWD.OPENFB]) OTE(MC_N255[98].10) ,XIC(MC_CIP_AV07.CW.[CWD.CLOSEDFB]) OTE(MC_N255[98].11) ,XIC(MC_CIP_AV07.CW.[CWD.FAULT]) OTE(MC_N255[98].15) ];
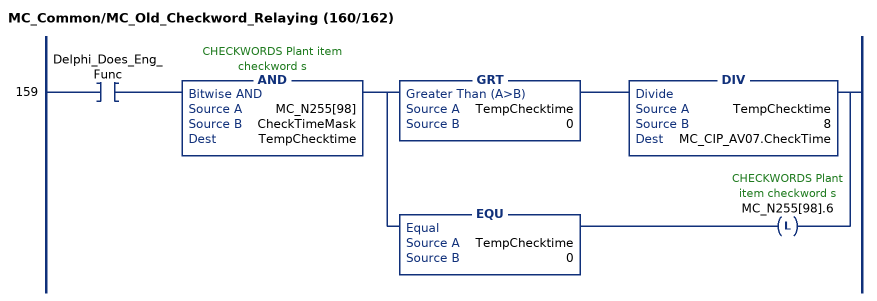
   159: XIC(Delphi_Does_Eng_Func)AND(MC_N255[98],CheckTimeMask,TempChecktime)[GRT(TempChecktime,0) DIV(TempChecktime,8,MC_CIP_AV07.CheckTime) ,EQU(TempChecktime,0) OTL(MC_N255[98].6) ];
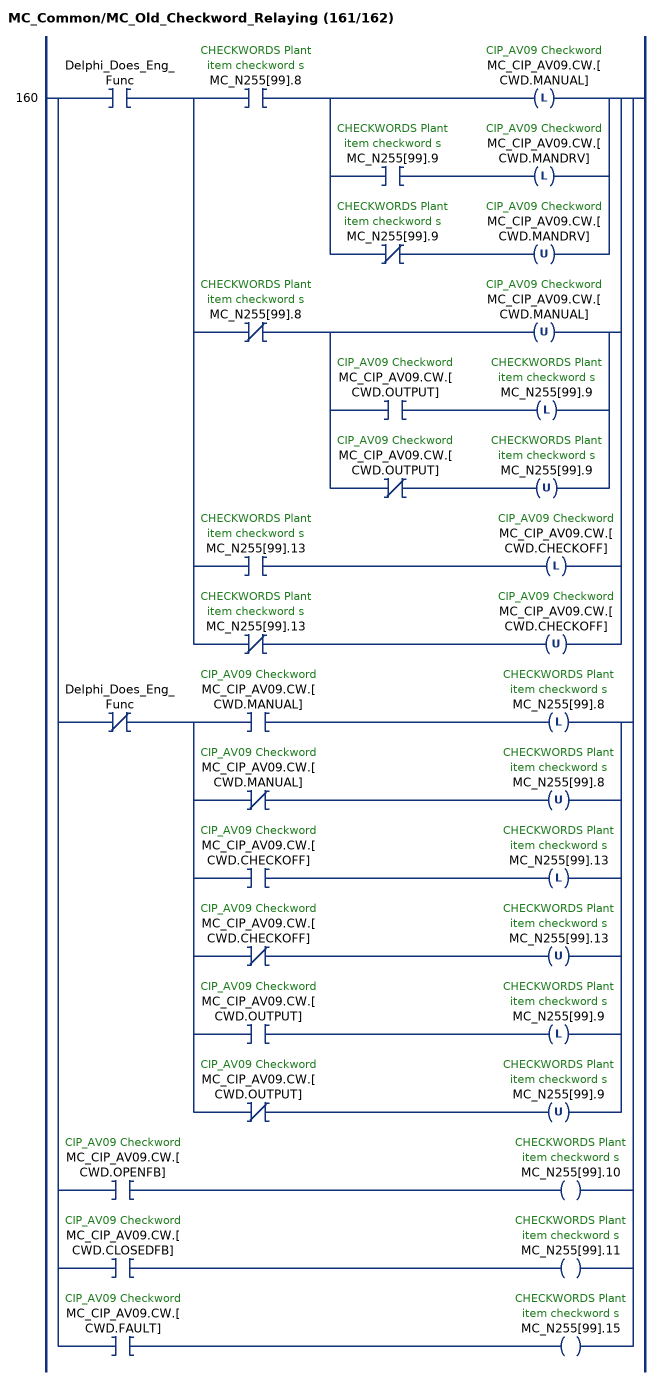
   160: [XIC(Delphi_Does_Eng_Func) [[XIC(MC_N255[99].8) [OTL(MC_CIP_AV09.CW.[CWD.MANUAL]) ,XIC(MC_N255[99].9) OTL(MC_CIP_AV09.CW.[CWD.MANDRV]) ,XIO(MC_N255[99].9) OTU(MC_CIP_AV09.CW.[CWD.MANDRV]) ] ,XIO(MC_N255[99].8) [OTU(MC_CIP_AV09.CW.[CWD.MANUAL]) ,[XIC(MC_CIP_AV09.CW.[CWD.OUTPUT]) OTL(MC_N255[99].9) ,XIO(MC_CIP_AV09.CW.[CWD.OUTPUT]) OTU(MC_N255[99].9) ] ] ] ,[XIC(MC_N255[99].13) OTL(MC_CIP_AV09.CW.[CWD.CHECKOFF]) ,XIO(MC_N255[99].13) OTU(MC_CIP_AV09.CW.[CWD.CHECKOFF]) ] ] ,XIO(Delphi_Does_Eng_Func) [[XIC(MC_CIP_AV09.CW.[CWD.MANUAL]) OTL(MC_N255[99].8) ,XIO(MC_CIP_AV09.CW.[CWD.MANUAL]) OTU(MC_N255[99].8) ] ,[XIC(MC_CIP_AV09.CW.[CWD.CHECKOFF]) OTL(MC_N255[99].13) ,XIO(MC_CIP_AV09.CW.[CWD.CHECKOFF]) OTU(MC_N255[99].13) ] ,[XIC(MC_CIP_AV09.CW.[CWD.OUTPUT]) OTL(MC_N255[99].9) ,XIO(MC_CIP_AV09.CW.[CWD.OUTPUT]) OTU(MC_N255[99].9) ] ] ,XIC(MC_CIP_AV09.CW.[CWD.OPENFB]) OTE(MC_N255[99].10) ,XIC(MC_CIP_AV09.CW.[CWD.CLOSEDFB]) OTE(MC_N255[99].11) ,XIC(MC_CIP_AV09.CW.[CWD.FAULT]) OTE(MC_N255[99].15) ];
